// Mitsubishi GX Works2 project: 30国轩预化成10.29,排队位置优化   PLC: Q10UDEH (continued)
	
			IF NOT ConveyorIO30134.xEmpty THEN(*有料时，旋转，转到2旋转完成*)
				ConveyorIO30134.xUnloadCCW:=ComConveyorIO30111.i_iResponsPCPLC=4;
				MOV(ComConveyorIO30111.i_iResponsPCPLC=4,2, RotorIO30401.iDestinationPos);(*4是左排，5是右排。左排转，右排不转*)
				MOV(ComConveyorIO30111.i_iResponsPCPLC=5,1, RotorIO30401.iDestinationPos);				
				IF (ComConveyorIO30111.i_iResponsPCPLC=4 AND  RotorIO30401.iCurrentPos=2 AND X61 )(*需要转，则等转到位置2,*)
					OR (ComConveyorIO30111.i_iResponsPCPLC=5 AND  RotorIO30401.iCurrentPos=1 AND X60 ) THEN(*不转则位置1为完成*)
					m_xRotor30401Done:=1;
				ELSE
						m_xRotor30401Done:=0;	
				END_IF;	
			ELSE(*无料就旋转回去，复位完成信号*)
				RotorIO30401.iDestinationPos:=1;
					m_xRotor30401Done:=0;
			END_IF;	
	(*预化成1入库转台下料*)		
	ConveyorIO30134.xUnload:=ConveyorIO30112.xEmpty 
														AND m_xRotor30401Done
														AND LifterIO30215.iCurrentPos=1 AND X5D;(*升降气缸*)
	ConveyorIO30112.xLoad:=ConveyorIO30134.xNextRun;
	IF ldp(TRUE,ConveyorIO30134.diDesConveyorOut>0) THEN
		ConveyorIO30112.diDesConveyorIn:=ConveyorIO30134.diDesConveyorOut;
		ConveyorIO30112.iTaskIDIn:=ConveyorIO30134.iTaskIDOut;
		ConveyorIO30112.iProductCategoryIn:=ConveyorIO30134.iProductCategoryOut;
	END_IF;
	(*预化成1入库气缸顶起*)
	LifterIO30215.xMDIExe:=NOT ConveyorIO30112.xError AND NOT ConveyorIO30112.xBusy;
	IF NOT ConveyorIO30112.xEmpty THEN
		LifterIO30215.iDestinationPos:=2;
	ELSE
		LifterIO30215.iDestinationPos:=1;
	END_IF;		
(***********************1巷道出库转台处理，运到转台上*********************)
	(*预化成1出库升降台控制*)
		IF ConveyorIO30114.xEmpty (*出库这里的开关位置要更改，改高点，不然putinto信号刷不到*)
			AND NOT ConveyorIO30114.xCWPresent
			AND NOT ConveyorIO30114.xCCWPresent
			AND NOT ConveyorIO30114.xBusy THEN
				LifterIO30214.iDestinationPos:=2;	
		ELSIF NOT ConveyorIO30114.xEmpty THEN
				LifterIO30214.iDestinationPos:=1;
		END_IF;	
			LifterIO30214.xMDIExe:=NOT ConveyorIO30114.xError AND NOT ConveyorIO30133.xError;
			DMOVP(ComConveyorIO30114.i_iResponsPCPLC=4,4,ConveyorIO30114.diDesConveyor);(*【需不需要转台转的信号生成】*)
			DMOVP(ComConveyorIO30114.i_iResponsPCPLC=5,5,ConveyorIO30114.diDesConveyor);(*【需不需要转台转的信号生成】*)			
			ConveyorIO30133.diDesConveyorIn:=ConveyorIO30114.diDesConveyorOut;(*【传递给转台】*)
			ConveyorIO30114.xUnload:=LifterIO30214.iCurrentPos=1 AND X5B(*升降台放下来*)
																	AND RotorIO30402.iCurrentPos=1 AND X62(*转台在接料位*)
																	 AND ConveyorIO30133.xEmpty(*转台为空*)
																	 AND ComConveyor30114.o_xReqSuccess(*旋转信号接收成功*);
			ConveyorIO30133.xLoad:=ConveyorIO30114.xNextRun;
	(*预化成1出库转台旋转控制*)		
		RotorIO30402.xMDIExe:=NOT ConveyorIO30133.xError AND NOT ConveyorIO30114.xError;
			IF NOT ConveyorIO30133.xEmpty THEN(*有料时，旋转，转到2旋转完成*)
				ConveyorIO30133.xUnloadCCW:=ConveyorIO30133.diDesConveyor=4;
				MOV(ConveyorIO30133.diDesConveyor=4,2, RotorIO30402.iDestinationPos);
				MOV(ConveyorIO30133.diDesConveyor=5,1, RotorIO30402.iDestinationPos);				
				IF (ConveyorIO30133.diDesConveyor=4 AND  RotorIO30402.iCurrentPos=2 AND X63 )(*需要转，则等转到位置2,*)
					OR (ConveyorIO30133.diDesConveyor=5 AND  RotorIO30402.iCurrentPos=1 AND X62 ) THEN(*不转则位置1为完成*)
					m_xRotor30402Done:=1;
				ELSE
					m_xRotor30402Done:=0;	
				END_IF;	
			ELSE(*无料就旋转回去，复位完成信号*)
				RotorIO30402.iDestinationPos:=1;
				m_xRotor30402Done:=0;
			END_IF;		
	(*化成1出库转台下料*)
		ConveyorIO30133.xUnload:=ConveyorIO30113.xEmpty 
														AND m_xRotor30402Done
														AND m_iTask30306=2;(*出库任务*)
(***********************1巷道出库的抢占任务，一边是产品出口，一边是2巷道的料路过*********************)	
	Task30306(xCondition:= Task30306Condition,
						xTaskComplete:= LDP(TRUE,ConveyorIO30110.xEmpty ),
	 					xReset:=g_xResetSingle AND g_diDeviceIDSelect=30110,
						 iPriority:=m_iTask30306);
		Task30306Condition[2]:=NOT ConveyorIO30133.xEmpty AND  m_xRotor30402Done ;(*正常出库*)(*这里需要等待旋转完成信号*)
		Task30306Condition[1]:=NOT ConveyorIO30106.xEmpty AND  ConveyorIO30106.diDesConveyor=30116;(*2巷道的入库要料*)
		DMOV(m_iTask30306=2, 30121, ConveyorIO30113.diDesConveyor );
	(*以上是1巷道出库顶升移载的抢占任务*)
	SwitchIO30306.xEntryEnable:=ConveyorIO30133.xNextRun;
	SwitchIO30306.xSwithEnable:=1;
	SwitchIO30306.xExitEnable:=ConveyorIO30138.xEmpty;
	(*任务1,去2巷道任务*)
	IF m_iTask30306=1 THEN
		IF ConveyorIO30110.xEmpty THEN
			SwitchIO30306.xLiftCylinderExtend:=0;
			SwitchIO30306.xLiftCylinderRetract:=1;
		ELSIF LDP(TRUE,NOT ConveyorIO30110.xEmpty) THEN
			SwitchIO30306.xLiftCylinderExtend:=1;
			SwitchIO30306.xLiftCylinderRetract:=0;	
		END_IF;
		ConveyorIO30110.xLoad:=ConveyorIO30106.xNextRun;
		ConveyorIO30110.diDesConveyorIn:=ConveyorIO30106.diDesConveyorOut;
		DMOVP(NOT ConveyorIO30110.xEmpty,ConveyorIO30106.diDesConveyor,ConveyorIO30113.diDesConveyor);(*【switch只能把目标地址传给入conveyor，不然会被写成0】*)
		SET(LDP(TRUE,NOT ConveyorIO30110.xEmpty) AND ConveyorIO30113.xEmpty,ConveyorIO30113.xPutInto);(*这里只要putinto了，就会进入switch正常流程了*)
		RST(LDP(TRUE,NOT ConveyorIO30113.xEmpty),ConveyorIO30113.xPutInto);	
	END_IF;
	(*任务为2时，顶升先升一下*)
	IF LDP(TRUE,m_iTask30306=2) THEN
			SwitchIO30306.xLiftCylinderExtend:=1;
			SwitchIO30306.xLiftCylinderRetract:=0;
		END_IF;	
	(*后续运给2巷道入库顶升移载*)
	ConveyorIO30138.diDesConveyorIn:=ConveyorIO30110.diDesConveyorOut;(*【目标地址传给138】*)
	ConveyorIO30138.xLoad:=ConveyorIO30110.xNextRun;
	ConveyorIO30138.xUnload:=ConveyorIO30115.xEmpty;
	ConveyorIO30115.diDesConveyorIn:=ConveyorIO30138.diDesConveyorOut;(*【目标地址传到2巷道顶升移载】*)
	SwitchIO30307.xEntryEnable:=ConveyorIO30138.xNextRun;
	SwitchIO30307.xSwithEnable:=ConveyorIO30115.diDesConveyor=30116;
	SwitchIO30307.xExitEnable:=(SwitchIO30307.xSwithEnable AND m_xLocation2Empty)(*需要转到2库，则2这边空就下料*)
															OR (NOT SwitchIO30307.xSwithEnable AND ConveyorIO30115.diDesConveyor=30121
																	AND m_iTask30308=2 AND ConveyorIO30122.xEmpty);(*不需要转，则等顶升移载308生成2任务*)
	m_xLocation2Load:=ConveyorIO30116.xNextRun;
(**************************************2巷道旋转，入库处理*****************************************************)
	(*定位机发出料请求，我要把门升起来，再给他发下料信号*)
	LifterIO30205.xMDIExe:=NOT ConveyorIO30132.xError;
		IF m_xLocation2NextRun AND ConveyorIO30132.xEmpty THEN
			LifterIO30205.iDestinationPos:=2;
		ELSE 
			LifterIO30205.iDestinationPos:=1;
		END_IF;	
	(*预化成2入库转台上料*)		
		m_xLocation2Unload:= ConveyorIO30132.xEmpty AND m_xLocation2NextRun(*他有下料请求时，我才判断*)
														AND RotorIO30403.iCurrentPos=1 AND X65(*转台在位置1才上料*)
														(*AND  LifterIO30205.iCurrentPos=2 AND X33*);												
		ConveyorIO30132.xLoad:=m_xLocation2NextRun 
															 AND RotorIO30403.iCurrentPos=1 AND X65
															(*AND  LifterIO30205.iCurrentPos=2 AND X33*) ;
	(*预化成2入库旋转控制*)		
		RotorIO30403.xMDIExe:=NOT ConveyorIO30132.xError AND NOT ConveyorIO30117.xError;
	
			IF NOT ConveyorIO30132.xEmpty THEN(*有料时，旋转，转到2旋转完成*)
				ConveyorIO30132.xUnloadCCW:=ComConveyorIO30116.i_iResponsPCPLC=4;
				MOV(ComConveyorIO30116.i_iResponsPCPLC=4,2, RotorIO30403.iDestinationPos);(*4是左排，5是右排。左排转，右排不转*)
				MOV(ComConveyorIO30116.i_iResponsPCPLC=5,1, RotorIO30403.iDestinationPos);				
				IF (ComConveyorIO30116.i_iResponsPCPLC=4 AND  RotorIO30403.iCurrentPos=2 AND X64 )(*需要转，则等转到位置2,*)
					OR (ComConveyorIO30116.i_iResponsPCPLC=5 AND  RotorIO30403.iCurrentPos=1 AND X65) THEN(*不转则位置1为完成*)
					m_xRotor30403Done:=1;
				ELSE
						m_xRotor30403Done:=0;	
				END_IF;	
			ELSE(*无料就旋转回去，复位完成信号*)
				RotorIO30403.iDestinationPos:=1;
					m_xRotor30403Done:=0;
			END_IF;	
(*预化成2入库转台下料*)		
	ConveyorIO30132.xUnload:=ConveyorIO30117.xEmpty 
														AND m_xRotor30403Done
														AND LifterIO30213.iCurrentPos=1 AND X59;(*升降气缸*)
	ConveyorIO30117.xLoad:=ConveyorIO30132.xNextRun;
	IF ldp(TRUE,ConveyorIO30132.diDesConveyorOut>0) THEN
		ConveyorIO30117.diDesConveyorIn:=ConveyorIO30132.diDesConveyorOut;
		ConveyorIO30117.iTaskIDIn:=ConveyorIO30132.iTaskIDOut;
		ConveyorIO30117.iProductCategoryIn:=ConveyorIO30132.iProductCategoryOut;
	END_IF;
	(*预化成2入库气缸顶起*)
	LifterIO30213.xMDIExe:=NOT ConveyorIO30117.xError AND NOT ConveyorIO30117.xBusy;
	IF NOT ConveyorIO30117.xEmpty THEN
		LifterIO30213.iDestinationPos:=2;
	ELSE
		LifterIO30213.iDestinationPos:=1;
	END_IF;		
(***********************2巷道出库转台处理，运到转台上*********************)
	(*预化成2出库升降台控制*)
		IF ConveyorIO30119.xEmpty (*出库这里的开关位置要更改，改高点，不然putinto信号刷不到*)
			AND NOT ConveyorIO30119.xCWPresent
			AND NOT ConveyorIO30119.xCCWPresent
			AND NOT ConveyorIO30119.xBusy THEN
				LifterIO30212.iDestinationPos:=2;	
		ELSIF NOT ConveyorIO30119.xEmpty THEN
				LifterIO30212.iDestinationPos:=1;
		END_IF;	
			LifterIO30212.xMDIExe:=NOT ConveyorIO30119.xError AND NOT ConveyorIO30131.xError;
			DMOVP(ComConveyorIO30119.i_iResponsPCPLC=4,4,ConveyorIO30119.diDesConveyor);(*【需不需要转台转的信号生成】*)
			DMOVP(ComConveyorIO30119.i_iResponsPCPLC=5,5,ConveyorIO30119.diDesConveyor);(*【需不需要转台转的信号生成】*)			
			ConveyorIO30131.diDesConveyorIn:=ConveyorIO30119.diDesConveyorOut;(*【传递给转台】*)
			ConveyorIO30119.xUnload:=LifterIO30212.iCurrentPos=1 AND X57(*升降台放下来*)
																	AND RotorIO30404.iCurrentPos=1 AND X66(*转台在接料位*)
																	 AND ConveyorIO30131.xEmpty(*转台为空*)
																	 AND ComConveyor30119.o_xReqSuccess(*旋转信号接收成功*);
			ConveyorIO30131.xLoad:=ConveyorIO30119.xNextRun;
(*预化成2出库旋转控制*)		
		RotorIO30404.xMDIExe:=NOT ConveyorIO30131.xError AND NOT ConveyorIO30119.xError;
			IF NOT ConveyorIO30131.xEmpty THEN(*有料时，旋转，转到2旋转完成*)
				ConveyorIO30131.xUnloadCCW:=ConveyorIO30131.diDesConveyor=4;
				MOV(ConveyorIO30131.diDesConveyor=4,2, RotorIO30404.iDestinationPos);
				MOV(ConveyorIO30131.diDesConveyor=5,1, RotorIO30404.iDestinationPos);				
				IF (ConveyorIO30131.diDesConveyor=4 AND  RotorIO30404.iCurrentPos=2 AND X67 )(*需要转，则等转到位置2,*)
					OR (ConveyorIO30131.diDesConveyor=5 AND  RotorIO30404.iCurrentPos=1 AND X66 ) THEN(*不转则位置1为完成*)
					m_xRotor30404Done:=1;
				ELSE
					m_xRotor30404Done:=0;	
				END_IF;	
			ELSE(*无料就旋转回去，复位完成信号*)
				RotorIO30404.iDestinationPos:=1;
				m_xRotor30404Done:=0;
			END_IF;		
(*化成2出库转台下料*)
		ConveyorIO30131.xUnload:=ConveyorIO30118.xEmpty 
														AND m_xRotor30404Done
														AND m_iTask30308=1;(*出库任务*)

(***********************2巷道出库的抢占任务，一边是产品出口，一边是1巷道出料路过*********************)	
	Task30308(xCondition:= Task30308Condition,
						xTaskComplete:= LDP(TRUE,ConveyorIO30121.xEmpty),
	 					xReset:=g_xResetSingle AND g_diDeviceIDSelect=30122,
						 iPriority:=m_iTask30308);
		Task30308Condition[1]:=NOT ConveyorIO30131.xEmpty AND m_xRotor30404Done ;(*正常出库*)
		Task30308Condition[2]:=NOT ConveyorIO30115.xEmpty AND  ConveyorIO30115.diDesConveyor<>30116;(*横向来料*)
	(*以上是2巷道出库顶升移载的抢占任务*)
	(*2巷道出库顶升移载任务1---2巷道出库任务*)
	SwitchIO30308.xEntryEnable:=ConveyorIO30131.xNextRun;
	SwitchIO30308.xSwithEnable:=1;
	SwitchIO30308.xExitEnable:=ConveyorIO30121.xEmpty;(*分拣那边有料时，这边不下料，防止赌住*)

	(*2巷道出库顶升移载任务2---1巷道的出料任务*)	
	IF m_iTask30308=2 THEN
		IF ConveyorIO30122.xEmpty THEN
			SwitchIO30308.xLiftCylinderExtend:=0;
			SwitchIO30308.xLiftCylinderRetract:=1;
		ELSIF LDP(TRUE,NOT ConveyorIO30122.xEmpty) THEN
			SwitchIO30306.xLiftCylinderExtend:=1;
			SwitchIO30306.xLiftCylinderRetract:=0;		
		END_IF;
		ConveyorIO30122.xLoad:=ConveyorIO30115.xNextRun;
		SET(LDP(TRUE,NOT ConveyorIO30122.xEmpty),ConveyorIO30118.xPutInto);(*这里只要putinto了，就会进入switch正常流程了*)
		RST(LDP(TRUE,NOT ConveyorIO30118.xEmpty),ConveyorIO30118.xPutInto);	
	END_IF;
	IF LDP(TRUE,m_iTask30306=1) THEN
			SwitchIO30308.xLiftCylinderExtend:=1;
			SwitchIO30308.xLiftCylinderRetract:=0;
		END_IF;	
	ConveyorIO30121.xLoad:=ConveyorIO30122.xNextRun;
	Y245:=D421.4 OR (g_xManual AND M594);	(*阻挡控制*)
	out_t(D421.4, TC3 , k30 );(**这里先留点时间给阻挡，再下料*)
	ConveyorIO30121.xUnload:=TS3 AND D421.5;
	D221.4:=ConveyorIO30121.xNextRun;
(*分拣完成信号控制*)(*
IF g_xPickOver AND NOT ConveyorIO30121.xEmpty THEN
	g_xPickDone:=1;
ELS*)IF 	ConveyorIO30121.xEmpty THEN 
	g_xPickDone:=0;	
END_IF;	

(**下层控制*)
D221.6:=ConveyorIO30124.xEmpty;
ConveyorIO30124.xLoad:=D421.6;
ConveyorIO30124.xUnload:=ConveyorIO30125.xEmpty;
ConveyorIO30125.xLoad:=ConveyorIO30124.xNextRun;
ConveyorIO30125.xUnload:=ConveyorIO30126.xEmpty;
ConveyorIO30126.xLoad:=ConveyorIO30125.xNextRun;
ConveyorIO30126.xUnload:=ConveyorIO30130.xEmpty	 AND D401.0;
ConveyorIO30130.xLoad:=ConveyorIO30126.xNextRun;
ConveyorIO30130.xUnload:=D401.0;
D201.0:=ConveyorIO30130.xNextRun;



END_IF;(*g_xauto那个if*)
(*这个是给40那边的信号，因为不良品和扫码位合成一个了*)
(*D221.5:=ConveyorIO30122.xNextRun;*)(*扫码位Load*)(*现在又屏蔽了，走putinto流程*)
D221.7:=X1E AND g_xPickDone;(*扫码位光电*)
D221.9:=g_xPickDone AND X4;(*putinto信号*)(*这里改为参数写入完成，允许下料了，就putinto*)
IF NOT g_xAuto THEN
	D201.0:=0;
	D221.6:=0;
END_IF;	


(*报警数据*)
g_xAlarm:=NOT g_xEStop 
					OR Conveyorio30104.xError
					OR Conveyorio30137.xError
					OR Conveyorio30109.xError
					OR Conveyorio30111.xError
					OR Conveyorio30116.xError
					OR Conveyorio30134.xError
					OR Conveyorio30133.xError
					OR ConveyorIO30132.xError
					OR Conveyorio30131.xError
					OR Conveyorio30112.xError
					OR Conveyorio30114.xError
					OR Conveyorio30117.xError
					OR Conveyorio30119.xError
					OR Conveyorio30124.xError
					OR Conveyorio30125.xError
					OR ConveyorIO30126.xError
					OR Conveyorio30130.xError
					OR Conveyorio30134.xError
					OR RotorIO30401.xOvertimeAlarm					
					OR RotorIO30402.xOvertimeAlarm
					OR RotorIO30403.xOvertimeAlarm
					OR RotorIO30404.xOvertimeAlarm
					OR ComConveyorIO30103.i_iResponsPCPLC=101(*高温库扫码失败*)
					OR ComConveyorIO30111.i_iResponsPCPLC=101(*预化成1扫码失败*)
					OR ComConveyorIO30116.i_iResponsPCPLC=101(*预化成2扫码失败*)
					
					
					
					;
END_PROGRAM

FUNCTION_BLOCK ConveyorOld
VAR
  m_xPresentDelay : BOOL;  (* 有无判断延时 *)
  m_xLoadDelayOut : BOOL;  (* 上料延时输出 *)
  m_xInitial : BOOL;  (* 初始化 *)
  m_tUnloadTimer : TIME;  (* 下料计时器 *)
  m_tPresentDelayCurrentTime : TIME;
  m_tonUnloadAlam : TON;  (* 下料报警定时器 *)
  m_tonPresentDelay : TON;  (* 物料有无判断延时，防止误动作 *)
  m_tonNotArriveAlarm : TON;  (* 未到达报警计时 *)
  m_tonLoadDelay : TON;  (* 上料延时 *)
  m_tNotArriveCurrentTime : TIME;  (* 未到达报警计时当前时间 *)
  m_tLoadTimer : TIME;  (* 上料计时器 *)
  iStep : INT;  (* 上料步骤 *)
  m_wStateWord : INT;
END_VAR
VAR_IN_OUT
  ConveyorMotor : ConveyorIO;  (* 输送线输入输出 *)
END_VAR
VAR
  m_tonZoneClear : TON;  (* 初始化清除 *)
  m_tZoneClearCurrentTime : TIME;  (* 初始化清除当前时间 *)
  m_xAutoClear : BOOL;  (* 初始化清除标志位 *)
  m_xZoneClearDone : BOOL;  (* 初始化清除完成 *)
END_VAR
(*////////////////////////////////////////////////////////////////////////////////////////////////////////////
//传输线控制FB块，可控制单方向线体，双向旋转线体，支持双向上下料            
//线体初始化后为空的情况下输入xLoad信号即可进行上料动作，使用xLoadCCW信号可反方向上料
//增加了产品信息和产品种类的储存，当传输线为空和上料进行标志位为零的情况下清除产品信息和产品种类
//使用方式是在置位xLoad信号后，把产品信息和产品种类传入，等下料后自动清零
//线体不为空的情况下使用xUnload信号可进行下料动作，物料有无传感器的下降沿后出发计时器，延时断开传输线旋转
//单方向传输线体把xLoadCCW、xUnloadCCW设置为零，双向线体上料方向和下料反向的,方向固定的 把xUnloadCCW设置为1
//双方向线体双向都能上下料的要根据上料的方向来设置xLoadCCW,xUnloadCCW
//增加工作中信号xBusy当电机正转 显示为工作中
//增加上下料超时报警，xLoadAlarm，xUnloadAlarm，设定时间在LOAD_UNLOAD_TIME常量上，现在设置的为30秒
//增加xPutInto信号，用于直接投入的物料，检测开关感应到后，直接进入下料流程，上升沿有效
//离开延时改为变量 iLeaveDelay 默认为0 离开检测开关离输送线尾端比较远的线体需要根据情况设定100ms为单位
//增加初始化标志位，增加进入延时时间，初始化为进入延时时间为0 ，离开延时时间为2S，通过外围接口可以更改
//修改信息  修改后请增加版本
//12-17进行了优化，增加了未到达报警，当物料未传送到下一设备，就报未到达报警，使用xNextRun标志位制作，没有正常到达
//第0步，不能跳转到第一步把标志位复位，即出现中断情况，2秒后报警
//修改信息  修改后请增加版本
上料延时增加为50ms防止干扰信号
nextrun信号在 第三步也要复位
增加限位报警
增加超宽报警
增加产品型号输出在下料的时候把产品型号输送给下一段线体
增加线体单独复位
增加任务插入功能配合全局变量
增加暂停功能
增加线体状态字显示  0 空闲 1：有料  2 工作中  3  超限报警 4 超宽报警  5 未到达报警  6 下料超时报警
空料判断放在自动前，进行有无报警判断，然后跳转
修改超限报警，与尺寸检测报警
初始化清除线体标志位xZoneClear
ZPA zero pressure accumulation  Term that describes the Conveyor controls and mechanical scheme that will 
cause loads to queue on a conveyor in discrete zones such that loads do not touch each other(wrapped boxed tray tote carton)
//YAO      V1.0
///////////////////////////////////////////////////////////////////////////////////////////////////////////
(*********************************************************)
(*//初始化，
//上料延时位0S，下料报警延时为30S
//下料延时设一个比较大的时间，主要依靠xunload标志位来停止输送线，特殊情况可以用延时来停止物流线下料
//设置时间大的时候计时器会失效*)
IF NOT m_xInitial THEN
	ConveyorMotor.tLoadDelay:=T#100ms;
	ConveyorMotor.tUnloadAlarmDelay:=T#30s;
	ConveyorMotor.xPosLimit:=1;
	ConveyorMotor.xNegLimit:=1;
	ConveyorMotor.xSizeDeficientDetect:=0;
	ConveyorMotor.xZoneClear:=0;
	ConveyorMotor.tZoneClearTime:=T#10s;
	m_xInitial:=1;
END_IF;
(*//自动
//复位信号把步号置0，但xLoad与xUnload没有复位，调用程序需要注意复位后把这两个信号置零，以免发生误动作
//物料有无判断增加延时，防止开自动瞬间误动作发生*)
m_tonPresentDelay(IN:= ConveyorMotor.xCWPresent OR ConveyorMotor.xCCWPresent,
                  PT:=T#100ms,
				  Q:= m_xPresentDelay,
				  ET:= m_tPresentDelayCurrentTime);

CASE iStep OF
	0:(*//初始化*)
	ConveyorMotor.xMotorCW:=0;
	ConveyorMotor.xMotorCCW:=0;
	ConveyorMotor.iProductCategoryOut:=0;
(*	//判断物料有无传感器*)	
		IF m_xPresentDelay THEN			
			ConveyorMotor.xEmpty:=0;
			IF g_xAuto AND NOT ConveyorMotor.xError THEN(*//自动情况下进行跳转*)(*无超限报警*)
				iStep:=3;
			END_IF;
		ELSE
			ConveyorMotor.xEmpty:=1;
			IF g_xAuto AND NOT ConveyorMotor.xError THEN(*//自动情况下进行跳转*)(*无超限报警*)
				iStep:=1;	
			END_IF;		
	END_IF;	
	1: (*//上料*)
	ConveyorMotor.xNextRun:=0;
	IF ConveyorMotor.xLoad    THEN (*//上料开始*)
		ConveyorMotor.iProductCategory:=0;	(*//上料开始清除产品信息*)
		iStep:=2;		
	END_IF;
	2: (*//上料完成*)
	IF ConveyorMotor.iProductCategoryIn<>0 THEN
		ConveyorMotor.iProductCategory:=ConveyorMotor.iProductCategoryIn;(* //产品信息传入*)
	END_IF;
	IF ConveyorMotor.xloadCCW THEN
		ConveyorMotor.xMotorCCW:=1; 
		ConveyorMotor.xMotorCW:=0;
	ELSE
	    ConveyorMotor.xMotorCW:=1;  
		ConveyorMotor.xMotorCCW:=0;
	END_IF;
		m_tonLoadDelay(IN:= (ConveyorMotor.xCWPresent AND NOT ConveyorMotor.xloadCCW) 
		                                        OR (ConveyorMotor.xCCWPresent AND ConveyorMotor.xloadCCW) ,
		                               PT:= ConveyorMotor.tLoadDelay ,
		                               Q:= m_xLoadDelayOut ,
		                               ET:= m_tLoadTimer );
	    IF m_xLoadDelayOut THEN 	 
		    iStep:=3;
		END_IF;
	3:(*//下料请求*)	
	ConveyorMotor.xMotorCW:=0;
	ConveyorMotor.xMotorCCW:=0;
	ConveyorMotor.xEmpty:=0;
	IF ConveyorMotor.xUnload AND NOT ConveyorMotor.xOverWidthAlarm  THEN (*无超宽报警可以下料*)
		iStep:=4;
	END_IF;
	4:(*	//下料完成*)
	IF ConveyorMotor.xUnloadCCW THEN   
		ConveyorMotor.xMotorCCW:=1;  
		ConveyorMotor.xMotorCW:=0;
		ELSE
	    ConveyorMotor.xMotorCW:=1;  
		ConveyorMotor.xMotorCCW:=0;
	END_IF;
	ConveyorMotor.xNextRun:=1; (*下一段线体旋转*)
	ConveyorMotor.iProductCategoryOut:=ConveyorMotor.iProductCategory;(*产品型号输出给下一段线体*)
	IF NOT ConveyorMotor.xUnload THEN 
		istep:=0;
	END_IF;
END_CASE;
(*In-feed zone clear and ready to accept a load from Upstream Conveyor*)
IF ldp(TRUE,g_xAuto) THEN
	m_xAutoClear:=1;
END_IF;
IF ldf(TRUE,g_xAuto) THEN
	m_xAutoClear:=0;
END_IF;
m_tonZoneClear(IN:= m_xAutoClear AND ConveyorMotor.xZoneClear ,PT:= ConveyorMotor.tZoneClearTime ,Q:=m_xZoneClearDone ,ET:= m_tZoneClearCurrentTime );
IF  m_xAutoClear AND ConveyorMotor.xZoneClear THEN
		ConveyorMotor.xMotorCW:=1; 
		iStep:=0;
END_IF;
IF ldf(TRUE, m_xAutoClear )THEN
	ConveyorMotor.xMotorCW:=0; 
END_IF;
IF NOT m_xAutoClear OR m_xZoneClearDone OR m_xPresentDelay THEN
	 m_xAutoClear:=0;
END_IF;	 
(*投入上料，搬出下料，也可用来初始化*)
IF LDP(TRUE,ConveyorMotor.xPutInto) THEN
	iStep:=0;
END_IF;
(*//当前任务显示*)
IF LDP(TRUE,ConveyorMotor.iDeviceID=g_iDeviceIDSelect) THEN
	g_iInsertTask:=ConveyorMotor.iProductCategory;
END_IF;
	(*//插入任务*)
IF g_xInsertTask AND ConveyorMotor.iDeviceID=g_iDeviceIDSelect THEN
	ConveyorMotor.iProductCategory:=g_iInsertTask;
END_IF;
(*//单线体复位，当设备号与本线体一致的时候执行复位*)
IF (g_xResetSingle AND ConveyorMotor.iDeviceID=g_iDeviceIDSelect)THEN (* //非正常情况下切断xNextRun不会复位，通过这个标志位会出发报警*)(*增加单体复位*)
	iStep:=0;
	ConveyorMotor.xNextRun:=0; 
	ConveyorMotor.xLimitAlarrm:=0;
	ConveyorMotor.xOverWidthAlarm:=0;
END_IF;
(*//手动*)
IF g_xManual THEN
(*	iStep:=0; *)(*//手动后上下料程序步骤清零*)
	(*//正转*)
	IF ConveyorMotor.xForward 
		AND ConveyorMotor.xBackward=0 
		AND ConveyorMotor.xMotorCCW=0 
		AND g_xEStop THEN
		ConveyorMotor.xMotorCW:=1;
		ConveyorMotor.xMotorCCW:=0;
		ELSE
		ConveyorMotor.xMotorCW:=0;
	END_IF;
	(*//反转*)
	IF ConveyorMotor.xBackward 
		AND ConveyorMotor.xForward=0 
		AND ConveyorMotor.xMotorCW=0 
		AND g_xEStop THEN
		ConveyorMotor.xMotorCCW:=1;
		conveyormotor.xMotorCW:=0;
		ELSE
		ConveyorMotor.xMotorCCW:=0;
	END_IF;
END_IF;
(*暂停*)
IF g_xPause THEN
	ConveyorMotor.xMotorCCW:=0;
	ConveyorMotor.xMotorCW:=0;
END_IF;
(*工作中信号输出*)
ConveyorMotor.xBusy:=ConveyorMotor.xMotorCCW OR ConveyorMotor.xMotorCW;
(*//未到达报警*)
m_tonNotArriveAlarm(IN:= iStep=0 AND ConveyorMotor.xNextRun  ,PT:= T#2s,Q:= ConveyorMotor.xNotArriveAlarm ,ET:= m_tNotArriveCurrentTime );
(*//下料超时报警*)
m_tonUnloadAlam(IN:= iStep=4,PT:=ConveyorMotor.tUnloadAlarmDelay,Q:= ConveyorMotor.xUnloadAlarm,ET:=m_tUnloadTimer );
(*//限位报警,进料检测开关失效*)
IF ( ((ConveyorMotor.xloadCCW AND NOT ConveyorMotor.xNegLimit)            (*反转上料，碰到负限位*)
	OR  ( NOT ConveyorMotor.xloadCCW AND NOT ConveyorMotor.xPosLimit)) (*正转上料，碰到正限位*)
    AND iStep=2) (*上料过程*)
    OR
   ( iStep=4 (*下料过程*)
	AND( (ConveyorMotor.xUnloadCCW AND NOT ConveyorMotor.xPosLimit)  
	OR (NOT ConveyorMotor.xUnloadCCW AND NOT ConveyorMotor.xNegLimit)))    
    THEN
    ConveyorMotor.xLimitAlarrm:=1;
    iStep:=0;
END_IF;
(*//超宽报警*)
IF (iStep=3 OR iStep=1) AND (NOT ConveyorMotor.xNegLimit OR NOT ConveyorMotor.xPosLimit) THEN
	ConveyorMotor.xOverWidthAlarm:=1;
END_IF;
(*//尺寸不足报警*)
(*//有料状态下检测两个开关都要有信号*)
IF iStep=3 AND ConveyorMotor.xSizeDeficientDetect AND (NOT ConveyorMotor.xCCWPresent OR NOT ConveyorMotor.xCWPresent)  THEN
	   ConveyorMotor.xOverWidthAlarm:=1;
	    iStep:=0;               
END_IF;
(*//总报警*)
ConveyorMotor.xError:=ConveyorMotor.xLimitAlarrm
                                              OR ConveyorMotor.xNotArriveAlarm
                                              OR ConveyorMotor.xUnloadAlarm                                             
                                              OR ConveyorMotor.xOverWidthAlarm;

(*//状态输出*)(*状态显示，容易造成指针容量不足*)
IF ConveyorMotor.xEmpty AND NOT ConveyorMotor.xBusy THEN
	m_wStateWord:=0;
END_IF;
IF ConveyorMotor.xEmpty=0 THEN
		m_wStateWord:=1;
END_IF;
IF ConveyorMotor.xBusy THEN
		m_wStateWord:=2;
END_IF;
IF ConveyorMotor.xLimitAlarrm THEN
		m_wStateWord:=3;
END_IF;
IF ConveyorMotor.xOverWidthAlarm THEN
		m_wStateWord:=4;
END_IF;
IF ConveyorMotor.xNotArriveAlarm THEN	
		m_wStateWord:=5;
END_IF;
IF ConveyorMotor.xUnloadAlarm THEN
		m_wStateWord:=6;	
END_IF;
(*选择本线体后，将状态赋值给全局变量进行显示*)
IF ConveyorMotor.iDeviceID=g_iDeviceIDSelect THEN
	g_iConveyorStatus:=m_wStateWord;
END_IF;
END_FUNCTION_BLOCK

FUNCTION_BLOCK ShuttleCar
VAR_IN_OUT
  ShuttleCarInOut : ShuttleCarIO;
END_VAR
VAR
  m_tonBrakeDelay : TON;  (* 延时 *)
  m_tBrakeDelayCurrentTime : TIME;
  m_tonArriveDelay : TON;  (* 到达延时计时器 *)
  m_xArriveDelay : BOOL;  (* 到达延时 *)
  m_tArriveDelayCurrentTime : TIME;  (* 到达延时当前时间 *)
  m_xInit : BOOL;  (* 初始化标志位 *)
  m_tonPauseDelay : TON;  (* 暂停减速 *)
  m_tPauseDelayCurrentTime : TIME;  (* 暂停延时当前时间 *)
  m_tonOvertimeAlarm : TON;  (* 超时报警定时器 *)
  m_tOvertimeCurrentTime : TIME;  (* 超时报警当前时间 *)
END_VAR
(*******************************************************************
输送小车程序，可用于使用认址片控制位置的输送车程序，可用于控制提升机，
使用了限位捕捉程序防止小车惯性过大冲过限位后继续行走，捕捉程序采用反
转复位，这样设计有弊端可能反转复位后车的位置并没有回到限位以内,当两个
限位同时碰到的时候，会使运料小车进入死锁状态，通过xPassLimit来解开死锁，
可以在触摸屏中使用一个带权限的按钮来进行控制，配合ShuttleCarCurrentPos
函数来计算位置信息
增加自动开始后将当前位置置为零的信号防止设备停在两个位置开关的中间
修改信息  修改后请增加版本
2018-1-22增加到位延时：到位延时时间可以设置，适应双向到位的位置开关，通过调整延时时间让穿梭车停在到位开关的中间
增加气缸控制信号 ShuttleCarInOut.xCylinder
增加抱闸延时 ShuttleCarInOut.tBrakeDelay
增加超时报警 ShuttleCarInOut.xOvertimeAlarm
YAO      V1.0
2018-1-22 YAO V1.1
2018-6-3：增加点动xMoveStep，单体报警复位
接口说明：
输入：
xReady    准备就绪信号，接变频器的准备就绪，无准备就绪信号的设备常置1
xForward   手动 正转
xBackward 手动 反转
iCurrentPos 当前位置信息，由外部函数给出
iDestinationPos  目标位置，自动情况下判断目标位置和当前位置的差，选择前进或后退
xPosLimit 正方向限位  常闭信号
xNegLimit 反方向限位  常闭信号
xMDIExe   自动行走使能
xPassLimit 限位屏蔽
tArriveDelay 到位延时时间设置，当前位置等于目标位置后延时相应时间后停止，默认为0
xCylinder 如果是气缸的把这个标志位置为1，
tBrakeDelay 打开抱闸延时，默认100ms。行走后会延时相应的时间打开抱闸，防止提升轴的掉落
xLooseDetect 松绳检测开关
输出：
xCW 正转输出
xCCW 反转输出
xBrake 抱闸输出 
xMDIDone 自动行走完成信号
xPosLimitCatch 正限位报警
xNegLimitCatch 负限位报警
xBusy 工作中信号
xLooseAlarm 松绳报警，报警后不可以下降，提升后如果没有松绳检测开关后复位报警信号


********************************************************************)
IF NOT m_xInit THEN
	ShuttleCarInOut.tArriveDelay:=T#0s;   (*到位延时初始化为0*)
	ShuttleCarInOut.tBrakeDelay:=T#100ms;(*抱闸延时初始化为100ms*)
	ShuttleCarInOut.tSetOverTime:=T#60s;(*超时报警初始化为1分钟*)
	m_xInit:=1;
END_IF;
(*如果是气缸的话屏蔽限位和Ready信号*)
IF ShuttleCarInOut.xCylinder THEN
	ShuttleCarInOut.xPosLimit:=1;
	ShuttleCarInOut.xNegLimit:=1;
	ShuttleCarInOut.xReady:=1;
END_IF;
(*限位捕捉，防止冲过限位开关，反转后复位*)
ShuttleCarInOut.xPosLimitCatch:=LDF(TRUE,ShuttleCarInOut.xPosLimit) OR ShuttleCarInOut.xPosLimitCatch;
IF ShuttleCarInOut.xCCW THEN  
	ShuttleCarInOut.xPosLimitCatch:=0;
END_IF;

ShuttleCarInOut.xNegLimitCatch:=LDF(TRUE,ShuttleCarInOut.xNegLimit) OR ShuttleCarInOut.xNegLimitCatch;
(*松绳报警*)
IF LDP(TRUE,ShuttleCarInOut.xLooseDetect) THEN	
	ShuttleCarInOut.xLooseAlarm:=1;
END_IF;
(*提升复位报警*)
IF ShuttleCarInOut.xCW AND NOT  ShuttleCarInOut.xLooseDetect THEN   
	ShuttleCarInOut.xLooseAlarm:=0; 
END_IF;

IF ShuttleCarInOut.xCW THEN   
	ShuttleCarInOut.xNegLimitCatch:=0; 
END_IF;

IF ShuttleCarInOut.xPassLimit OR
	g_xReset OR   (*增加复位按钮*)
	(ShuttleCarInOut.xNegLimitCatch 
	AND ShuttleCarInOut.xPosLimitCatch)  THEN  
	ShuttleCarInOut.xNegLimitCatch:=0; 
	ShuttleCarInOut.xPosLimitCatch:=0;
	ShuttleCarInOut.xLooseAlarm:=0;
END_IF;
IF ShuttleCarInOut.xReady AND g_xEStop THEN
(*手动*)
    IF g_xManual THEN  
	    IF ShuttleCarInOut.xForward 
			AND ShuttleCarInOut.xBackward=0 
			AND ShuttleCarInOut.xCCW=0 
			AND ShuttleCarInOut.xPosLimitCatch=0  THEN
		    ShuttleCarInOut.xCW:=1;
		    ELSE
		    ShuttleCarInOut.xCW:=0;
	    END_IF;
	    IF ShuttleCarInOut.xBackward 
			AND ShuttleCarInOut.xForward=0 
			AND ShuttleCarInOut.xCW=0 
			AND ShuttleCarInOut.xNegLimitCatch=0 
			AND ShuttleCarInOut.xLooseAlarm=0
			AND G_xEStop THEN  
		    ShuttleCarInOut.xCCW:=1;
		    ELSE
		    ShuttleCarInOut.xCCW:=0;
	    END_IF;
    END_IF;
    (**********)
(*自动*)
  IF g_xAuto OR ShuttleCarInOut.xMoveStep   THEN  
  	(*点动*)
  	IF LDP(TRUE,ShuttleCarInOut.xMoveStep)  THEN (*点动模式后把当前位置赋值给目标位置，防止误动作*)
  		ShuttleCarInOut.iDestinationPos:=ShuttleCarInOut.iCurrentPos;
  		END_IF;
 		IF LDP(TRUE,ShuttleCarInOut.xForward) AND ShuttleCarInOut.xMoveStep THEN
 			ShuttleCarInOut.xMDIExe:=1;
			ShuttleCarInOut.iDestinationPos:=ShuttleCarInOut.iCurrentPos+1;
		END_IF;
		IF LDP(TRUE,ShuttleCarInOut.xBackward) AND ShuttleCarInOut.xMoveStep AND ShuttleCarInOut.iCurrentPos>0  THEN
			ShuttleCarInOut.xMDIExe:=1;
			ShuttleCarInOut.iDestinationPos:=ShuttleCarInOut.iCurrentPos-1;
		END_IF;	 
	(*>>>>>>>>>>>>>>>>>>>>>>>>>>>>>>>>>>>>>*)	
	  IF ShuttleCarInOut.xMDIExe AND ShuttleCarInOut.iDestinationPos<>0 THEN	
	    IF ShuttleCarInOut.iCurrentPos<ShuttleCarInOut.iDestinationPos AND ShuttleCarInOut.xPosLimitCatch=0 THEN   (*正转*)
			ShuttleCarInOut.xCW:=1;
			ShuttleCarInOut.xCCW:=0;
			ShuttleCarInOut.xMDIDone:=0;
		END_IF;

		IF ShuttleCarInOut.iCurrentPos>ShuttleCarInOut.iDestinationPos AND ShuttleCarInOut.xNegLimitCatch=0 AND ShuttleCarInOut.xLooseAlarm=0 THEN   (*反转*)
			ShuttleCarInOut.xCCW:=1;
			ShuttleCarInOut.xCW:=0;
			ShuttleCarInOut.xMDIDone:=0;
		END_IF;
	m_tonArriveDelay(IN:= ShuttleCarInOut.iCurrentPos=ShuttleCarInOut.iDestinationPos ,
	                                    PT:= ShuttleCarInOut.tArriveDelay ,
	                                    Q:= m_xArriveDelay ,
	                                    ET:= m_tArriveDelayCurrentTime);
	     (*到位延时时间可以设置，适应双向到位的位置开关，通过调整延时时间让穿梭车停在到位开关的中间*)
		IF m_xArriveDelay AND NOT ShuttleCarInOut.xCylinder THEN
			ShuttleCarInOut.xCW:=0;
			ShuttleCarInOut.xCCW:=0;
			ShuttleCarInOut.xMDIDone:=1;
			ELSE
			ShuttleCarInOut.xMDIDone:=0;
		END_IF;

		IF ShuttleCarInOut.xPosLimitCatch THEN
			ShuttleCarInOut.xCW:=0;
			ShuttleCarInOut.xMDIDone:=0;
		END_IF;

		IF ShuttleCarInOut.xNegLimitCatch  OR ShuttleCarInOut.xLooseAlarm THEN
			ShuttleCarInOut.xCCW:=0;
			ShuttleCarInOut.xMDIDone:=0;
		END_IF;
		ELSE
		ShuttleCarInOut.xCW:=0;
		ShuttleCarInOut.xCCW:=0;
		ShuttleCarInOut.xMDIDone:=0;
	  END_IF;
	END_IF;
	ELSE  (*无就绪信号   或急停的情况下*)
		ShuttleCarInOut.xCW:=0;
		ShuttleCarInOut.xCCW:=0;	
END_IF;
    (*抱闸延时*)
m_tonBrakeDelay(IN:= ShuttleCarInOut.xCW OR ShuttleCarInOut.xCCW,
                                    PT:= ShuttleCarInOut.tBrakeDelay,
                                    Q:=ShuttleCarInOut.xBrake ,
                                    ET:= m_tBrakeDelayCurrentTime);

(*自动上电后把当前位置清零，防止穿梭车不在开关位置*)
IF LDP(TRUE,g_xAuto) THEN
	ShuttleCarInOut.iCurrentPos:=0;
END_IF;
IF ShuttleCarInOut.xCW OR ShuttleCarInOut.xCCW THEN
	ShuttleCarInOut.xBusy:=1;
	ELSE
	ShuttleCarInout.xBusy:=0;
END_IF;

(*暂停，带延时减速斜坡，ShuttleCarInOut.xPauseRamp为减速斜坡输出位*)
m_tonPauseDelay(IN:=g_xPause,PT:= T#2s ,Q:=ShuttleCarInOut.xPauseRamp,ET:= m_tPauseDelayCurrentTime );
IF ShuttleCarInOut.xPauseRamp THEN
	ShuttleCarInOut.xCW:=0;
	ShuttleCarInOut.xCCW:=0;
	ShuttleCarInOut.xBrake:=0;
END_IF;
(*超时报警*)
m_tonOvertimeAlarm(IN:= ShuttleCarInOut.xMDIExe AND (ShuttleCarInOut.iCurrentPos<>ShuttleCarInOut.iDestinationPos) ,
                                           PT:= ShuttleCarInOut.tSetOverTime,
                                           Q:= ShuttleCarInOut.xOvertimeAlarm ,
                                           ET:= m_tOvertimeCurrentTime );
(*//单体复位，当设备号与本设备一致的时候执行复位*)
IF (g_xResetSingle AND ShuttleCarInOut.diDeviceID=g_diDeviceIDSelect)THEN(*增加单体复位*)
	ShuttleCarInOut.iCurrentPos:=0;
END_IF;
END_FUNCTION_BLOCK

FUNCTION_BLOCK Switch
VAR_IN_OUT
  ConveyorEntryIO : ConveyorIO;
  ConveyorExitIO : ConveyorIO;
END_VAR
VAR
  m_tonLiftCylinderDelay : TON;  (* 顶升延时 *)
  m_xLiftCylinderDelay : BOOL;
  m_tLiftCylinderDelay : TIME;
  m_tonExitBarDelay : TON;  (* 退出阻挡器延时 *)
  m_tExitBarDelay : TIME;
  m_xExitBarDelay : BOOL;
END_VAR
VAR_IN_OUT
  SwitchIO : SwitchIO;
END_VAR
VAR
  iStep : INT;
  m_xInitial : BOOL;
  m_tonCylinderOvertime : TON;  (* 气缸超时报警定时器 *)
  m_tCylinderOvertimeCurrent : TIME;
END_VAR
(**************************************************
//顶升移载模块，抽象为一条输入输线 ，一条输出输送线
//一个进入阻挡器，一个放出阻挡器，和一个顶升气缸的控制
//程序思路比较混乱，接口不清晰，需要整改
//直接放行的时候有问题
//switchEnable =0的时候   离开线体的PutInto有问题
//增加xPutInto程序
//12-17日   V1.0
//***************************************************)
(*ConveyorEntry(ConveyorMotor:=ConveyorEntryIO);
(*ConveyorExit(ConveyorMotor:=ConveyorExitIO);*)


IF NOT m_xInitial THEN
	SwitchIO.tSetOvertime:=T#5s;
	SwitchIO.xExitEnable:=1;
	m_xInitial:=1;
END_IF;
IF g_xAuto THEN
	CASE iStep OF
		0:(*初始化*)
		ConveyorEntryIO.xLoad:=0;
		ConveyorEntryIO.xUnload:=0;
		ConveyorEntryIO.xPutInto:=0;
		ConveyorExitIO.xLoad:=0;
		ConveyorExitIo.xUnload:=0;
		ConveyorExitIO.xPutInto:=0;
		SwitchIO.xEntryBarCylinderRetract:=0;
		SwitchIO.xExitBarCylinderRetract:=0;
		IF SwitchIO.xLiftCylinderExtendInit THEN
			SwitchIO.xLiftCylinderExtend:=1;
			SwitchIO.xLiftCylinderRetract:=0;
		    IF SwitchIO.xLiftCylinderExtendDetect THEN
			    iStep:=1;
			END_IF; 
			ELSE
			SwitchIO.xLiftCylinderExtend:=0;
			SwitchIO.xLiftCylinderRetract:=1;	
		    IF SwitchIO.xLiftCylinderRetractDetect THEN
			    iStep:=1;
		    END_IF;		
		END_IF;
		1:(*上料*)
        IF SwitchIO.xEntryEnable AND ConveyorEntryIO.xEmpty AND ConveyorExitIO.xEmpty THEN
        	SwitchIO.xEntryBarCylinderRetract:=1;
        	ConveyorEntryIO.xLoad:=1;
        END_IF;
        IF ConveyorEntryIO.xEmpty=0 THEN
        	SwitchIO.xEntryBarCylinderRetract:=0;
        	ConveyorEntryIO.xLoad:=0;
        	ConveyorExitIO.xPutInto:=ConveyorExitIO.xEmpty;
        END_IF;
        IF m_xLiftCylinderDelay AND  SwitchIO.xSwithEnable AND SwitchIO.xExitEnable THEN
			iStep:=2;
        END_IF;
        IF SwitchIO.xSwithEnable=0 AND m_xLiftCylinderDelay AND SwitchIO.xExitEnable  THEN
			iStep:=3;
        END_IF;
		2:(*顶升*)
		ConveyorExitIO.iProductCategory:=ConveyorEntryIO.iProductCategory;
		ConveyorExitIO.iTaskID:=ConveyorEntryIO.iTaskID;
		ConveyorExitIO.diDesConveyor:=ConveyorEntryIO.diDesConveyor;
		SwitchIO.xExitBarCylinderRetract:=0;
		ConveyorExitIO.xPutInto:=0;
		IF SwitchIO.xLiftCylinderExtendInit THEN
			SwitchIO.xLiftCylinderExtend:=0;
			SwitchIO.xLiftCylinderRetract:=1;
		    ELSE
			SwitchIO.xLiftCylinderExtend:=1;
			SwitchIO.xLiftCylinderRetract:=0;			
		END_IF;

		IF SwitchIO.xLiftCylinderExtendInit THEN
		  	IF SwitchIO.xLiftCylinderRetractDetect THEN
		  		iStep:=4;
		  	END_IF;
		  	ELSE
		  	IF SwitchIO.xLiftCylinderExtendDetect THEN
				iStep:=4; 
		  	END_IF;
		END_IF;
		3:(*放行*)	
		ConveyorExitIO.iProductCategory:=ConveyorEntryIO.iProductCategory;
		ConveyorExitIO.iTaskID:=ConveyorEntryIO.iTaskID;
		ConveyorExitIO.diDesConveyor:=ConveyorEntryIO.diDesConveyor;
		SwitchIO.xExitBarCylinderRetract:=1;
		ConveyorExitIO.xPutInto:=0;
		iStep:=4;
		4:(*下料*)
		(*通过出料传输线下料*)
		IF SwitchIO.xExitEnable  AND m_xExitBarDelay AND NOT SwitchIO.xExitBarCylinderRetract  THEN		  
		  	ConveyorExitIO.xUnload:=1;
			ELSE
		  	ConveyorExitIO.xUnload:=0;
		END_IF;	
		(*通过进料传输线下料*)
		IF SwitchIO.xExitEnable  AND m_xExitBarDelay  AND SwitchIO.xExitBarCylinderRetract THEN		  
		  	ConveyorEntryIO.xUnload:=1;
			ELSE
		  	ConveyorEntryIO.xUnload:=0;
		END_IF;			    	
		IF (ConveyorExitIO.xEmpty OR ConveyorEntryIO.xEmpty) AND m_xExitBarDelay  THEN
		  	ConveyorExitIO.xPutInto:=1;
		  	ConveyorEntryIO.xPutInto:=1;
			iStep:=0; 
		END_IF;
	END_CASE;
	m_tonLiftCylinderDelay(IN:=NOT ConveyorEntryIO.xEmpty AND iStep=1 ,PT:= T#1S ,Q:= m_xLiftCylinderDelay ,ET:=m_tLiftCylinderDelay );
	m_tonExitBarDelay(IN:=iStep=4 ,PT:= T#1s ,Q:= m_xExitBarDelay ,ET:= m_tExitBarDelay);
END_IF;
(*复位程序*)
IF (g_xResetSingle AND  (g_diDeviceIDSelect=ConveyorEntryIO.diDeviceID OR g_diDeviceIDSelect=ConveyorExitIO.diDeviceID))
	OR LDP(TRUE,SwitchIO.xLiftCylinderExtendInit) 
	OR LDF(TRUE,SwitchIO.xLiftCylinderExtendInit) 
	OR LDP(TRUE,SwitchIO.xPutInto)  THEN
	ConveyorEntryIO.xPutInto:=1;
	ConveyorExitIO.xPutInto:=1;
	iStep:=0;
END_IF;

IF g_xManual  THEN
	iStep:=0;
	ConveyorEntryIO.xLoad:=0;
    ConveyorEntryIO.xUnload:=0;
	ConveyorEntryIO.xPutInto:=0;
	ConveyorExitIO.xLoad:=0;
	ConveyorExitIo.xUnload:=0;
	ConveyorExitIO.xPutInto:=0;
	SwitchIO.xEntryBarCylinderRetract:=0;
	SwitchIO.xExitBarCylinderRetract:=0;
	IF SwitchIO.xEntryBarCylinderRetractButton THEN
		SwitchIO.xEntryBarCylinderRetract:=1;
		ELSE
		SwitchIO.xEntryBarCylinderRetract:=0;
	END_IF;
	IF SwitchIO.xExitBarCylinderRetractButton THEN
		SwitchIO.xExitBarCylinderRetract:=1;
		ELSE
		SwitchIO.xExitBarCylinderRetract:=0;
	END_IF;
	IF SwitchIO.xLiftCylinderExtendButton AND NOT SwitchIO.xLiftCylinderRetractButton THEN
		SwitchIO.xLiftCylinderExtend:=1;
		SwitchIO.xLiftCylinderRetract:=0;
	END_IF;
	IF NOT SwitchIO.xLiftCylinderExtendButton AND  SwitchIO.xLiftCylinderRetractButton THEN
		SwitchIO.xLiftCylinderExtend:=0;
		SwitchIO.xLiftCylinderRetract:=1;
	END_IF;		 
END_IF;
(*气缸超时报警*)
m_tonCylinderOvertime(IN:= (SwitchIO.xLiftCylinderExtend AND NOT SwitchIO.xLiftCylinderExtendDetect) 
OR  (SwitchIO.xLiftCylinderRetract AND NOT SwitchIO.xLiftCylinderRetractDetect) ,
PT:= SwitchIO.tSetOvertime ,Q:= SwitchIO.xOvertimeAlarm ,ET:= m_tCylinderOvertimeCurrent );
END_FUNCTION_BLOCK

